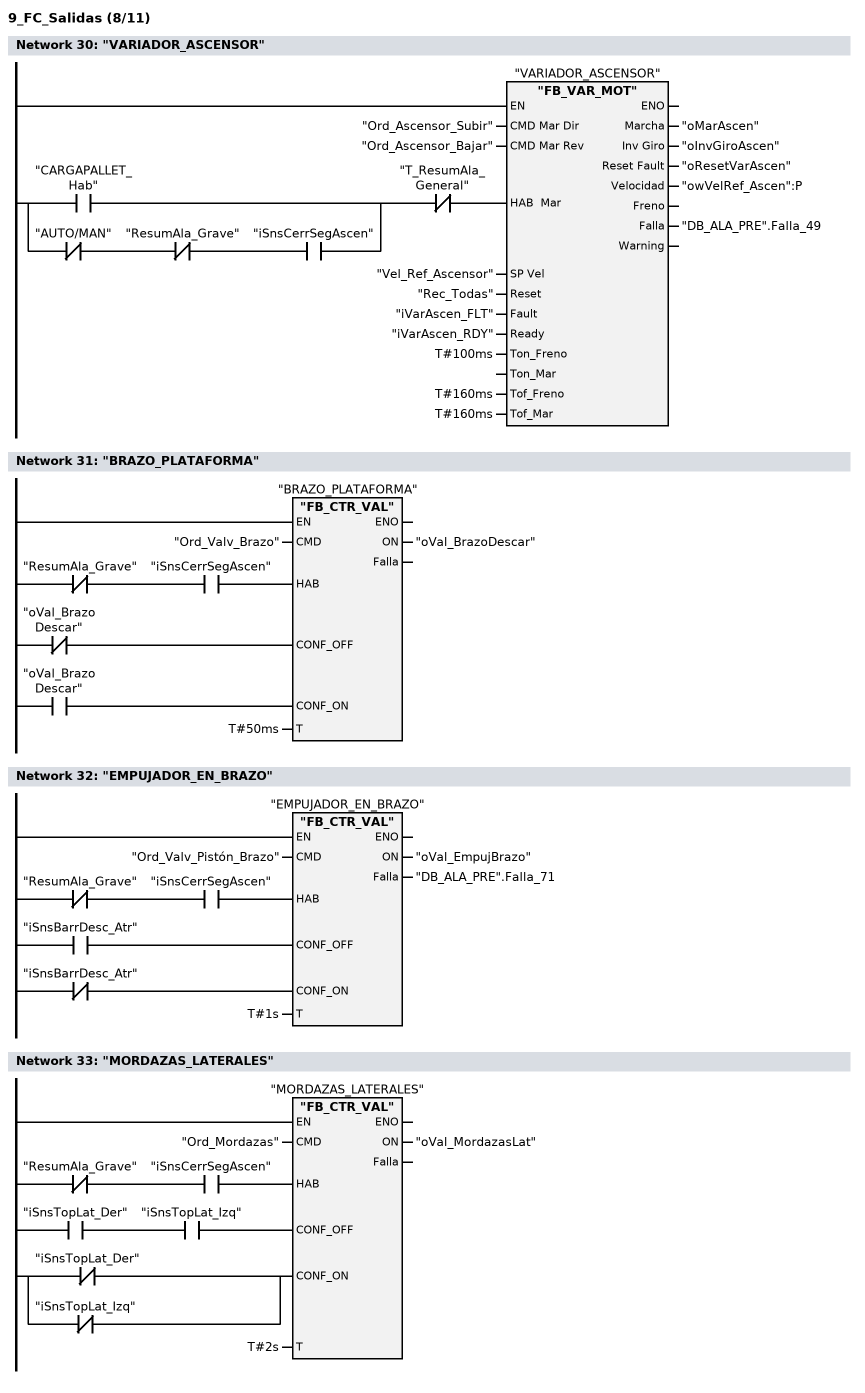
   RUNG wire#powerrail
      "VARIADOR_ASCENSOR"("HAB  Mar" := wire#w2, "CMD Mar Dir" := "Ord_Ascensor_Subir", "CMD Mar Rev" := "Ord_Ascensor_Bajar", "SP Vel" := "Vel_Ref_Ascensor", Reset := "Rec_Todas", Fault := "iVarAscen_FLT", Ready := "iVarAscen_RDY", Ton_Freno := T#100ms, Ton_Mar :=, Tof_Freno := T#160ms, Tof_Mar := T#160ms, Marcha => "oMarAscen", "Inv Giro" => "oInvGiroAscen", "Reset Fault" => "oResetVarAscen", Velocidad => "owVelRef_Ascen":P, Freno =>, Falla => "DB_ALA_PRE".Falla_49, Warning =>)
   END_RUNG
   RUNG wire#powerrail
      Contact( "CARGAPALLET_Hab" )
      wire#w1
      I_Contact( "T_ResumAla_General" )
   END_RUNG wire#w2
   RUNG wire#powerrail
      I_Contact( "AUTO/MAN" )
      I_Contact( "ResumAla_Grave" )
      Contact( "iSnsCerrSegAscen" )
   END_RUNG wire#w1
   // the same network as SCL:
   "VARIADOR_ASCENSOR"("CMD Mar Dir" := "Ord_Ascensor_Subir",   // "FB_VAR_MOT"
                       "CMD Mar Rev" := "Ord_Ascensor_Bajar",
                       "HAB  Mar" := ("CARGAPALLET_Hab" OR (NOT "AUTO/MAN" AND NOT "ResumAla_Grave" AND "iSnsCerrSegAscen")) AND NOT "T_ResumAla_General",
                       "SP Vel" := "Vel_Ref_Ascensor",
                       Reset := "Rec_Todas",
                       Fault := "iVarAscen_FLT",
                       Ready := "iVarAscen_RDY",
                       Ton_Freno := T#100ms,
                       Tof_Freno := T#160ms,
                       Tof_Mar := T#160ms,
                       Marcha => "oMarAscen",
                       "Inv Giro" => "oInvGiroAscen",
                       "Reset Fault" => "oResetVarAscen",
                       Velocidad => "owVelRef_Ascen":P,
                       Falla => "DB_ALA_PRE".Falla_49);
END_REGION

REGION Network 31: "BRAZO_PLATAFORMA"
   RUNG wire#powerrail
      "BRAZO_PLATAFORMA"(HAB := wire#w1, CONF_OFF := wire#w2, CONF_ON := wire#w3, CMD := "Ord_Valv_Brazo", T := T#50ms, ON => "oVal_BrazoDescar", Falla =>)
   END_RUNG
   RUNG wire#powerrail
      I_Contact( "ResumAla_Grave" )
      Contact( "iSnsCerrSegAscen" )
   END_RUNG wire#w1
   RUNG wire#powerrail
      I_Contact( "oVal_BrazoDescar" )
   END_RUNG wire#w2
   RUNG wire#powerrail
      Contact( "oVal_BrazoDescar" )
   END_RUNG wire#w3
   // the same network as SCL:
   "BRAZO_PLATAFORMA"(CMD := "Ord_Valv_Brazo",   // "FB_CTR_VAL"
                      HAB := NOT "ResumAla_Grave" AND "iSnsCerrSegAscen",
                      CONF_OFF := NOT "oVal_BrazoDescar",
                      CONF_ON := "oVal_BrazoDescar",
                      T := T#50ms,
                      ON => "oVal_BrazoDescar");
END_REGION

REGION Network 32: "EMPUJADOR_EN_BRAZO"
   RUNG wire#powerrail
      "EMPUJADOR_EN_BRAZO"(HAB := wire#w1, CONF_OFF := wire#w2, CONF_ON := wire#w3, CMD := "Ord_Valv_Pistón_Brazo", T := T#1s, ON => "oVal_EmpujBrazo", Falla => "DB_ALA_PRE".Falla_71)
   END_RUNG
   RUNG wire#powerrail
      I_Contact( "ResumAla_Grave" )
      Contact( "iSnsCerrSegAscen" )
   END_RUNG wire#w1
   RUNG wire#powerrail
      Contact( "iSnsBarrDesc_Atr" )
   END_RUNG wire#w2
   RUNG wire#powerrail
      I_Contact( "iSnsBarrDesc_Atr" )
   END_RUNG wire#w3
   // the same network as SCL:
   "EMPUJADOR_EN_BRAZO"(CMD := "Ord_Valv_Pistón_Brazo",   // "FB_CTR_VAL"
                        HAB := NOT "ResumAla_Grave" AND "iSnsCerrSegAscen",
                        CONF_OFF := "iSnsBarrDesc_Atr",
                        CONF_ON := NOT "iSnsBarrDesc_Atr",
                        T := T#1s,
                        ON => "oVal_EmpujBrazo",
                        Falla => "DB_ALA_PRE".Falla_71);
END_REGION

REGION Network 33: "MORDAZAS_LATERALES"
   RUNG wire#powerrail
      "MORDAZAS_LATERALES"(HAB := wire#w1, CONF_OFF := wire#w2, CONF_ON := wire#w3, CMD := "Ord_Mordazas", T := T#2s, ON => "oVal_MordazasLat", Falla =>)
   END_RUNG
   RUNG wire#powerrail
      I_Contact( "ResumAla_Grave" )
      Contact( "iSnsCerrSegAscen" )
   END_RUNG wire#w1
   RUNG wire#powerrail
      Contact( "iSnsTopLat_Der" )
      Contact( "iSnsTopLat_Izq" )
   END_RUNG wire#w2
   RUNG wire#powerrail
      I_Contact( "iSnsTopLat_Der" )
   END_RUNG wire#w3
   RUNG wire#powerrail
      I_Contact( "iSnsTopLat_Izq" )
   END_RUNG wire#w3
   // the same network as SCL:
   "MORDAZAS_LATERALES"(CMD := "Ord_Mordazas",   // "FB_CTR_VAL"
                        HAB := NOT "ResumAla_Grave" AND "iSnsCerrSegAscen",
                        CONF_OFF := "iSnsTopLat_Der" AND "iSnsTopLat_Izq",
                        CONF_ON := NOT "iSnsTopLat_Der" OR NOT "iSnsTopLat_Izq",
                        T := T#2s,
                        ON => "oVal_MordazasLat");
END_REGION

REGION Network 34: "MORDAZA_FINAL"
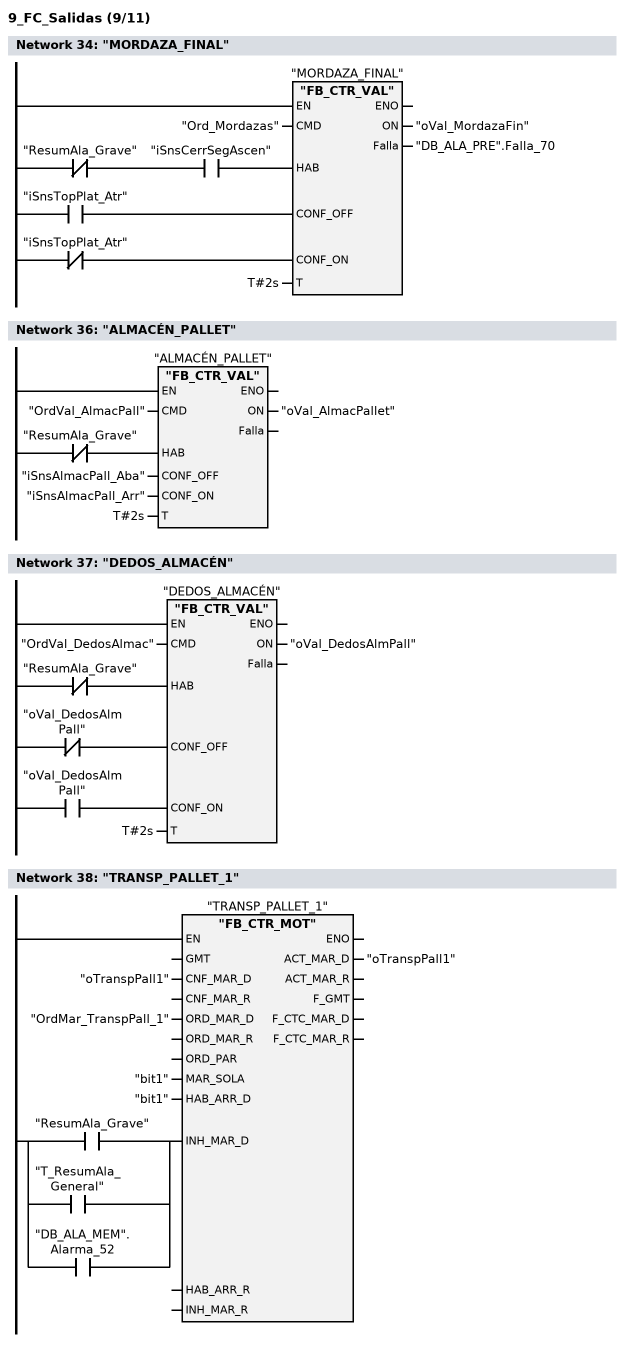
   RUNG wire#powerrail
      "MORDAZA_FINAL"(HAB := wire#w1, CONF_OFF := wire#w2, CONF_ON := wire#w3, CMD := "Ord_Mordazas", T := T#2s, ON => "oVal_MordazaFin", Falla => "DB_ALA_PRE".Falla_70)
   END_RUNG
   RUNG wire#powerrail
      I_Contact( "ResumAla_Grave" )
      Contact( "iSnsCerrSegAscen" )
   END_RUNG wire#w1
   RUNG wire#powerrail
      Contact( "iSnsTopPlat_Atr" )
   END_RUNG wire#w2
   RUNG wire#powerrail
      I_Contact( "iSnsTopPlat_Atr" )
   END_RUNG wire#w3
   // the same network as SCL:
   "MORDAZA_FINAL"(CMD := "Ord_Mordazas",   // "FB_CTR_VAL"
                   HAB := NOT "ResumAla_Grave" AND "iSnsCerrSegAscen",
                   CONF_OFF := "iSnsTopPlat_Atr",
                   CONF_ON := NOT "iSnsTopPlat_Atr",
                   T := T#2s,
                   ON => "oVal_MordazaFin",
                   Falla => "DB_ALA_PRE".Falla_70);
END_REGION

REGION Network 35: ----------------------------------------------------------------- TRANSPORTE DE PALLETS -----------------------------------------------------------------¬
END_REGION

REGION Network 36: "ALMACÉN_PALLET"
   RUNG wire#powerrail
      "ALMACÉN_PALLET"(HAB := wire#w1, CMD := "OrdVal_AlmacPall", CONF_OFF := "iSnsAlmacPall_Aba", CONF_ON := "iSnsAlmacPall_Arr", T := T#2s, ON => "oVal_AlmacPallet", Falla =>)
   END_RUNG
   RUNG wire#powerrail
      I_Contact( "ResumAla_Grave" )
   END_RUNG wire#w1
   // the same network as SCL:
   "ALMACÉN_PALLET"(CMD := "OrdVal_AlmacPall",   // "FB_CTR_VAL"
                    HAB := NOT "ResumAla_Grave",
                    CONF_OFF := "iSnsAlmacPall_Aba",
                    CONF_ON := "iSnsAlmacPall_Arr",
                    T := T#2s,
                    ON => "oVal_AlmacPallet");
END_REGION

REGION Network 37: "DEDOS_ALMACÉN"
   RUNG wire#powerrail
      "DEDOS_ALMACÉN"(HAB := wire#w1, CONF_OFF := wire#w2, CONF_ON := wire#w3, CMD := "OrdVal_DedosAlmac", T := T#2s, ON => "oVal_DedosAlmPall", Falla =>)
   END_RUNG
   RUNG wire#powerrail
      I_Contact( "ResumAla_Grave" )
   END_RUNG wire#w1
   RUNG wire#powerrail
      I_Contact( "oVal_DedosAlmPall" )
   END_RUNG wire#w2
   RUNG wire#powerrail
      Contact( "oVal_DedosAlmPall" )
   END_RUNG wire#w3
   // the same network as SCL:
   "DEDOS_ALMACÉN"(CMD := "OrdVal_DedosAlmac",   // "FB_CTR_VAL"
                   HAB := NOT "ResumAla_Grave",
                   CONF_OFF := NOT "oVal_DedosAlmPall",
                   CONF_ON := "oVal_DedosAlmPall",
                   T := T#2s,
                   ON => "oVal_DedosAlmPall");
END_REGION

REGION Network 38: "TRANSP_PALLET_1"
   RUNG wire#powerrail
      "TRANSP_PALLET_1"(INH_MAR_D := wire#w1, GMT :=, CNF_MAR_D := "oTranspPall1", CNF_MAR_R :=, ORD_MAR_D := "OrdMar_TranspPall_1", ORD_MAR_R :=, ORD_PAR :=, MAR_SOLA := "bit1", HAB_ARR_D := "bit1", HAB_ARR_R :=, INH_MAR_R :=, ACT_MAR_D => "oTranspPall1", ACT_MAR_R =>, F_GMT =>, F_CTC_MAR_D =>, F_CTC_MAR_R =>)
   END_RUNG
   RUNG wire#powerrail
      Contact( "ResumAla_Grave" )
   END_RUNG wire#w1
   RUNG wire#powerrail
      Contact( "T_ResumAla_General" )
   END_RUNG wire#w1
   RUNG wire#powerrail
      Contact( "DB_ALA_MEM".Alarma_52 )
   END_RUNG wire#w1
   // the same network as SCL:
   "TRANSP_PALLET_1"(CNF_MAR_D := "oTranspPall1",   // "FB_CTR_MOT"
                     ORD_MAR_D := "OrdMar_TranspPall_1",
                     MAR_SOLA := "bit1",
                     HAB_ARR_D := "bit1",
                     INH_MAR_D := "ResumAla_Grave" OR "T_ResumAla_General" OR "DB_ALA_MEM".Alarma_52,
                     ACT_MAR_D => "oTranspPall1");
END_REGION

REGION Network 39: "TRANSP_PALLET_2"
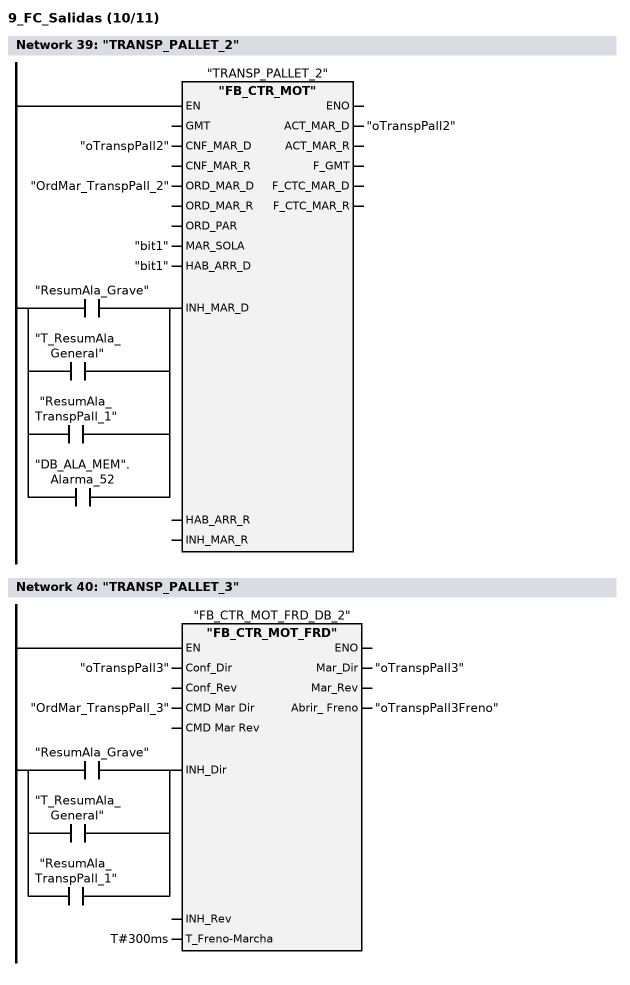
   RUNG wire#powerrail
      "TRANSP_PALLET_2"(INH_MAR_D := wire#w1, GMT :=, CNF_MAR_D := "oTranspPall2", CNF_MAR_R :=, ORD_MAR_D := "OrdMar_TranspPall_2", ORD_MAR_R :=, ORD_PAR :=, MAR_SOLA := "bit1", HAB_ARR_D := "bit1", HAB_ARR_R :=, INH_MAR_R :=, ACT_MAR_D => "oTranspPall2", ACT_MAR_R =>, F_GMT =>, F_CTC_MAR_D =>, F_CTC_MAR_R =>)
   END_RUNG
   RUNG wire#powerrail
      Contact( "ResumAla_Grave" )
   END_RUNG wire#w1
   RUNG wire#powerrail
      Contact( "T_ResumAla_General" )
   END_RUNG wire#w1
   RUNG wire#powerrail
      Contact( "ResumAla_TranspPall_1" )
   END_RUNG wire#w1
   RUNG wire#powerrail
      Contact( "DB_ALA_MEM".Alarma_52 )
   END_RUNG wire#w1
   // the same network as SCL:
   "TRANSP_PALLET_2"(CNF_MAR_D := "oTranspPall2",   // "FB_CTR_MOT"
                     ORD_MAR_D := "OrdMar_TranspPall_2",
                     MAR_SOLA := "bit1",
                     HAB_ARR_D := "bit1",
                     INH_MAR_D := "ResumAla_Grave" OR "T_ResumAla_General" OR "ResumAla_TranspPall_1" OR "DB_ALA_MEM".Alarma_52,
                     ACT_MAR_D => "oTranspPall2");
END_REGION

REGION Network 40: "TRANSP_PALLET_3"
   RUNG wire#powerrail
      "FB_CTR_MOT_FRD_DB_2"(INH_Dir := wire#w1, Conf_Dir := "oTranspPall3", Conf_Rev :=, "CMD Mar Dir" := "OrdMar_TranspPall_3", "CMD Mar Rev" :=, INH_Rev :=, "T_Freno-Marcha" := T#300ms, Mar_Dir => "oTranspPall3", Mar_Rev =>, "Abrir_ Freno" => "oTranspPall3Freno")
   END_RUNG
   RUNG wire#powerrail
      Contact( "ResumAla_Grave" )
   END_RUNG wire#w1
   RUNG wire#powerrail
      Contact( "T_ResumAla_General" )
   END_RUNG wire#w1
   RUNG wire#powerrail
      Contact( "ResumAla_TranspPall_1" )
   END_RUNG wire#w1
   // the same network as SCL:
   "FB_CTR_MOT_FRD_DB_2"(Conf_Dir := "oTranspPall3",   // "FB_CTR_MOT_FRD"
                         "CMD Mar Dir" := "OrdMar_TranspPall_3",
                         INH_Dir := "ResumAla_Grave" OR "T_ResumAla_General" OR "ResumAla_TranspPall_1",
                         "T_Freno-Marcha" := T#300ms,
                         Mar_Dir => "oTranspPall3",
                         "Abrir_ Freno" => "oTranspPall3Freno");
END_REGION

REGION Network 41: "TRANSP_PALLET_4"
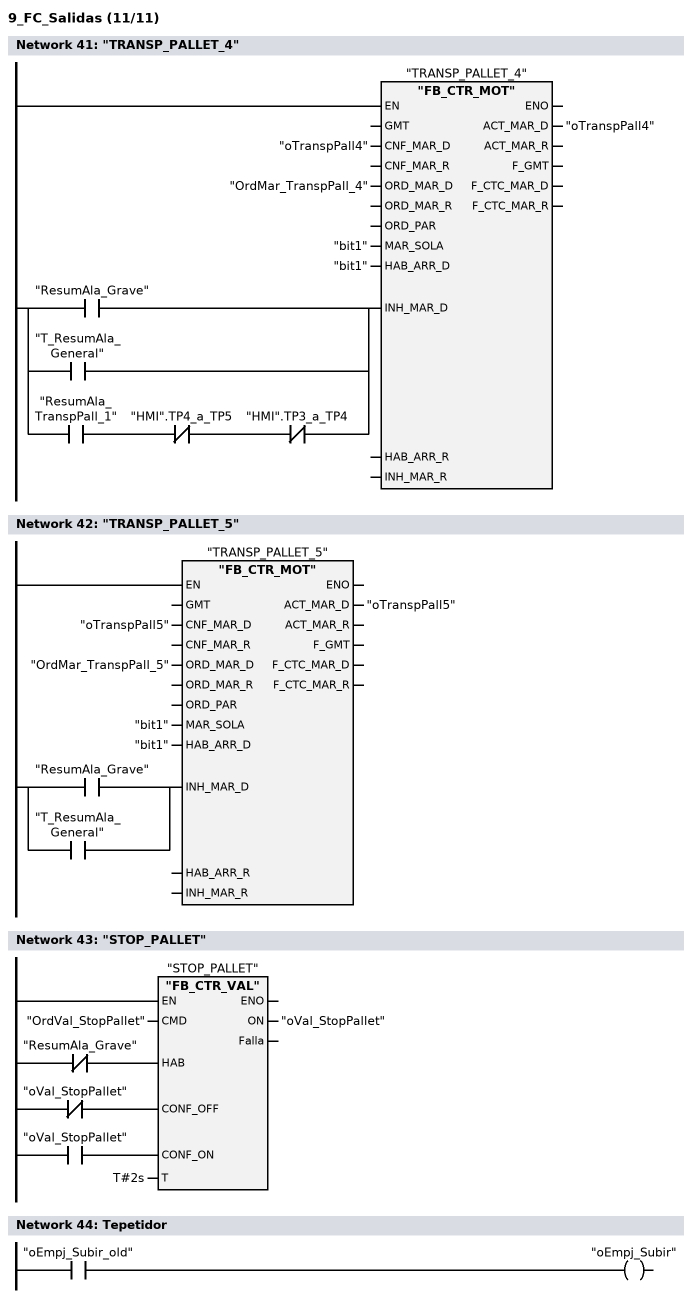
   RUNG wire#powerrail
      "TRANSP_PALLET_4"(INH_MAR_D := wire#w1, GMT :=, CNF_MAR_D := "oTranspPall4", CNF_MAR_R :=, ORD_MAR_D := "OrdMar_TranspPall_4", ORD_MAR_R :=, ORD_PAR :=, MAR_SOLA := "bit1", HAB_ARR_D := "bit1", HAB_ARR_R :=, INH_MAR_R :=, ACT_MAR_D => "oTranspPall4", ACT_MAR_R =>, F_GMT =>, F_CTC_MAR_D =>, F_CTC_MAR_R =>)
   END_RUNG
   RUNG wire#powerrail
      Contact( "ResumAla_Grave" )
   END_RUNG wire#w1
   RUNG wire#powerrail
      Contact( "T_ResumAla_General" )
   END_RUNG wire#w1
   RUNG wire#powerrail
      Contact( "ResumAla_TranspPall_1" )
      I_Contact( "HMI".TP4_a_TP5 )
      I_Contact( "HMI".TP3_a_TP4 )
   END_RUNG wire#w1
   // the same network as SCL:
   "TRANSP_PALLET_4"(CNF_MAR_D := "oTranspPall4",   // "FB_CTR_MOT"
                     ORD_MAR_D := "OrdMar_TranspPall_4",
                     MAR_SOLA := "bit1",
                     HAB_ARR_D := "bit1",
                     INH_MAR_D := "ResumAla_Grave" OR "T_ResumAla_General" OR ("ResumAla_TranspPall_1" AND NOT "HMI".TP4_a_TP5 AND NOT "HMI".TP3_a_TP4),
                     ACT_MAR_D => "oTranspPall4");
END_REGION

REGION Network 42: "TRANSP_PALLET_5"
   RUNG wire#powerrail
      "TRANSP_PALLET_5"(INH_MAR_D := wire#w1, GMT :=, CNF_MAR_D := "oTranspPall5", CNF_MAR_R :=, ORD_MAR_D := "OrdMar_TranspPall_5", ORD_MAR_R :=, ORD_PAR :=, MAR_SOLA := "bit1", HAB_ARR_D := "bit1", HAB_ARR_R :=, INH_MAR_R :=, ACT_MAR_D => "oTranspPall5", ACT_MAR_R =>, F_GMT =>, F_CTC_MAR_D =>, F_CTC_MAR_R =>)
   END_RUNG
   RUNG wire#powerrail
      Contact( "ResumAla_Grave" )
   END_RUNG wire#w1
   RUNG wire#powerrail
      Contact( "T_ResumAla_General" )
   END_RUNG wire#w1
   // the same network as SCL:
   "TRANSP_PALLET_5"(CNF_MAR_D := "oTranspPall5",   // "FB_CTR_MOT"
                     ORD_MAR_D := "OrdMar_TranspPall_5",
                     MAR_SOLA := "bit1",
                     HAB_ARR_D := "bit1",
                     INH_MAR_D := "ResumAla_Grave" OR "T_ResumAla_General",
                     ACT_MAR_D => "oTranspPall5");
END_REGION

REGION Network 43: "STOP_PALLET"
   RUNG wire#powerrail
      "STOP_PALLET"(HAB := wire#w1, CONF_OFF := wire#w2, CONF_ON := wire#w3, CMD := "OrdVal_StopPallet", T := T#2s, ON => "oVal_StopPallet", Falla =>)
   END_RUNG
   RUNG wire#powerrail
      I_Contact( "ResumAla_Grave" )
   END_RUNG wire#w1
   RUNG wire#powerrail
      I_Contact( "oVal_StopPallet" )
   END_RUNG wire#w2
   RUNG wire#powerrail
      Contact( "oVal_StopPallet" )
   END_RUNG wire#w3
   // the same network as SCL:
   "STOP_PALLET"(CMD := "OrdVal_StopPallet",   // "FB_CTR_VAL"
                 HAB := NOT "ResumAla_Grave",
                 CONF_OFF := NOT "oVal_StopPallet",
                 CONF_ON := "oVal_StopPallet",
                 T := T#2s,
                 ON => "oVal_StopPallet");
END_REGION

REGION Network 44: Tepetidor
   RUNG wire#powerrail
      Contact( "oEmpj_Subir_old" )
      Coil( "oEmpj_Subir" )
   END_RUNG
   // the same network as SCL:
   "oEmpj_Subir" := "oEmpj_Subir_old";
END_REGION
END_FUNCTION

FUNCTION "4_FC_Dosificador" : Void   // FC11, LAD
{ S7_Optimized_Access := 'FALSE' }
VERSION : 0.1
BEGIN

REGION Network 1: ESTADO ACTIVO
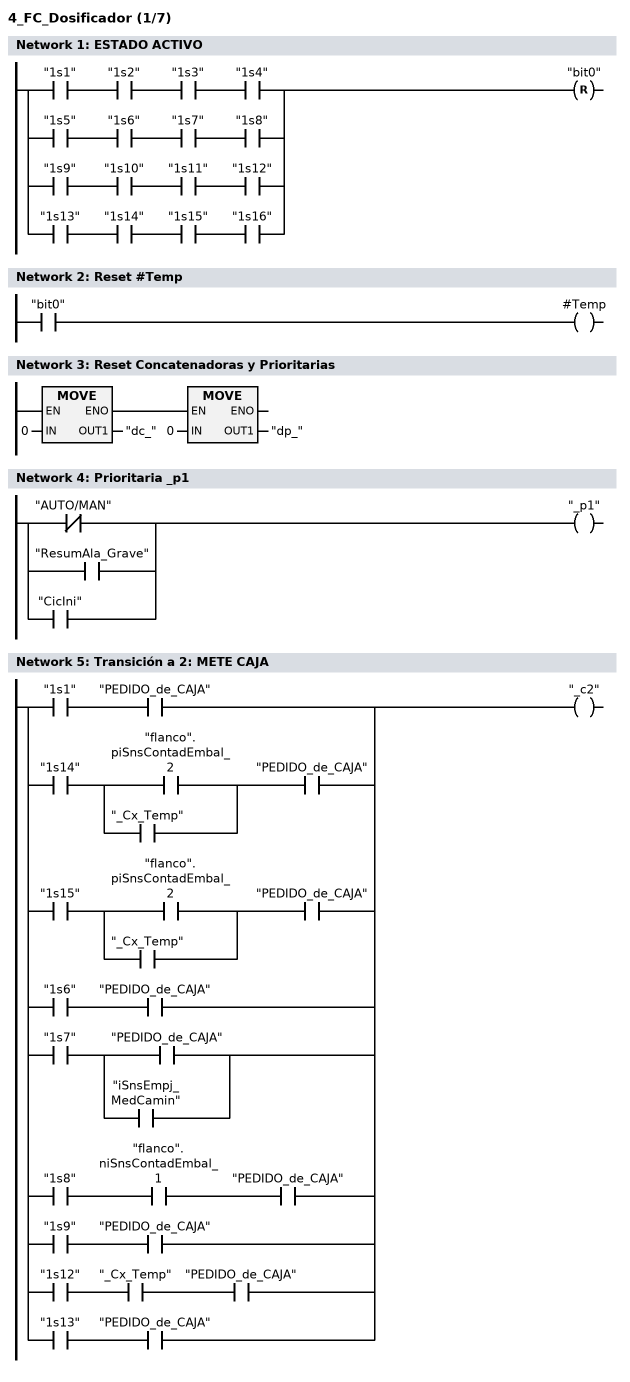
   RUNG wire#powerrail
      Contact( "1s1" )
      Contact( "1s2" )
      Contact( "1s3" )
      Contact( "1s4" )
      wire#w1
      R_Coil( "bit0" )
   END_RUNG
   RUNG wire#powerrail
      Contact( "1s5" )
      Contact( "1s6" )
      Contact( "1s7" )
      Contact( "1s8" )
   END_RUNG wire#w1
   RUNG wire#powerrail
      Contact( "1s9" )
      Contact( "1s10" )
      Contact( "1s11" )
      Contact( "1s12" )
   END_RUNG wire#w1
   RUNG wire#powerrail
      Contact( "1s13" )
      Contact( "1s14" )
      Contact( "1s15" )
      Contact( "1s16" )
   END_RUNG wire#w1
   // the same network as SCL:
   IF ("1s1" AND "1s2" AND "1s3" AND "1s4") OR ("1s5" AND "1s6" AND "1s7" AND "1s8") OR ("1s9" AND "1s10" AND "1s11" AND "1s12") OR ("1s13" AND "1s14" AND "1s15" AND "1s16") THEN
       "bit0" := FALSE;
   END_IF;
END_REGION

REGION Network 2: Reset #Temp
   RUNG wire#powerrail
      Contact( "bit0" )
      Coil( #Temp )
   END_RUNG
   // the same network as SCL:
   #Temp := "bit0";
END_REGION

REGION Network 3: Reset Concatenadoras y Prioritarias
   RUNG wire#powerrail
      { S7_GenerateENO := "TRUE" } Move(in := 0, out1 => "dc_")
      { S7_GenerateENO := "TRUE" } Move(in := 0, out1 => "dp_")
   END_RUNG
   // the same network as SCL:
   // ENO of a box is taken as its EN; it also drops when the box reports an error
   "dc_" := 0;
   "dp_" := 0;
END_REGION

REGION Network 4: Prioritaria _p1
   RUNG wire#powerrail
      I_Contact( "AUTO/MAN" )
      wire#w1
      Coil( "_p1" )
   END_RUNG
   RUNG wire#powerrail
      Contact( "ResumAla_Grave" )
   END_RUNG wire#w1
   RUNG wire#powerrail
      Contact( "CicIni" )
   END_RUNG wire#w1
   // the same network as SCL:
   "_p1" := NOT "AUTO/MAN" OR "ResumAla_Grave" OR "CicIni";
END_REGION

REGION Network 5: Transición a 2: METE CAJA
   RUNG wire#powerrail
      Contact( "1s1" )
      Contact( "PEDIDO_de_CAJA" )
      wire#w1
      Coil( "_c2" )
   END_RUNG
   RUNG wire#powerrail
      Contact( "1s14" )
      wire#w2
      Contact( "flanco".piSnsContadEmbal_2 )
      wire#w3
      Contact( "PEDIDO_de_CAJA" )
   END_RUNG wire#w1
   RUNG wire#w2
      Contact( "_Cx_Temp" )
   END_RUNG wire#w3
   RUNG wire#powerrail
      Contact( "1s15" )
      wire#w4
      Contact( "flanco".piSnsContadEmbal_2 )
      wire#w5
      Contact( "PEDIDO_de_CAJA" )
   END_RUNG wire#w1
   RUNG wire#w4
      Contact( "_Cx_Temp" )
   END_RUNG wire#w5
   RUNG wire#powerrail
      Contact( "1s6" )
      Contact( "PEDIDO_de_CAJA" )
   END_RUNG wire#w1
   RUNG wire#powerrail
      Contact( "1s7" )
      wire#w6
      Contact( "PEDIDO_de_CAJA" )
   END_RUNG wire#w1
   RUNG wire#w6
      Contact( "iSnsEmpj_MedCamin" )
   END_RUNG wire#w1
   RUNG wire#powerrail
      Contact( "1s8" )
      Contact( "flanco".niSnsContadEmbal_1 )
      Contact( "PEDIDO_de_CAJA" )
   END_RUNG wire#w1
   RUNG wire#powerrail
      Contact( "1s9" )
      Contact( "PEDIDO_de_CAJA" )
   END_RUNG wire#w1
   RUNG wire#powerrail
      Contact( "1s12" )
      Contact( "_Cx_Temp" )
      Contact( "PEDIDO_de_CAJA" )
   END_RUNG wire#w1
   RUNG wire#powerrail
      Contact( "1s13" )
      Contact( "PEDIDO_de_CAJA" )
   END_RUNG wire#w1
   // the same network as SCL:
   "_c2" := ("1s1" AND "PEDIDO_de_CAJA") OR ("1s14" AND ("flanco".piSnsContadEmbal_2 OR "_Cx_Temp") AND "PEDIDO_de_CAJA") OR ("1s15" AND ("flanco".piSnsContadEmbal_2 OR "_Cx_Temp") AND "PEDIDO_de_CAJA") OR ("1s6" AND "PEDIDO_de_CAJA") OR ("1s7" AND ("PEDIDO_de_CAJA" OR "iSnsEmpj_MedCamin")) OR ("1s8" AND "flanco".niSnsContadEmbal_1 AND "PEDIDO_de_CAJA") OR ("1s9" AND "PEDIDO_de_CAJA") OR ("1s12" AND "_Cx_Temp" AND "PEDIDO_de_CAJA") OR ("1s13" AND "PEDIDO_de_CAJA");
END_REGION

REGION Network 6: Transición a 3: FIGURA H
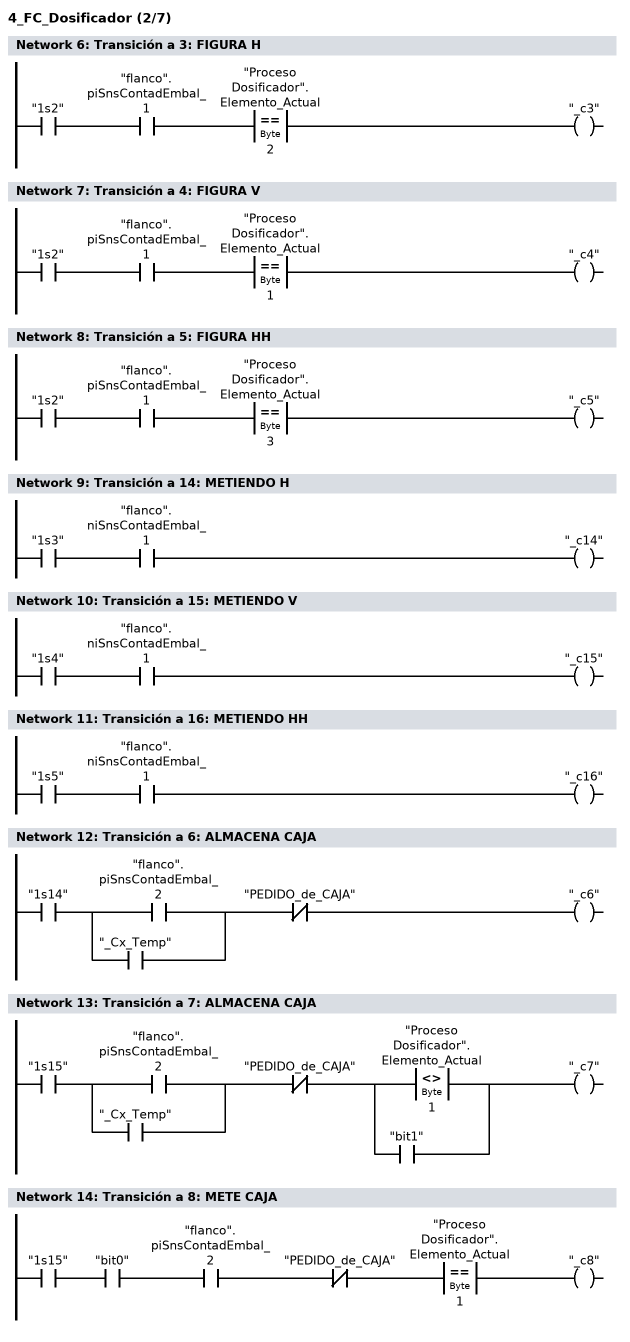
   RUNG wire#powerrail
      Contact( "1s2" )
      Contact( "flanco".piSnsContadEmbal_1 )
      { S7_Templates := "SrcType := Byte" } EQ_Contact(in1 := "Proceso Dosificador".Elemento_Actual, in2 := 2)
      Coil( "_c3" )
   END_RUNG
   // the same network as SCL:
   "_c3" := "1s2" AND "flanco".piSnsContadEmbal_1 AND ("Proceso Dosificador".Elemento_Actual = 2);
END_REGION

REGION Network 7: Transición a 4: FIGURA V
   RUNG wire#powerrail
      Contact( "1s2" )
      Contact( "flanco".piSnsContadEmbal_1 )
      { S7_Templates := "SrcType := Byte" } EQ_Contact(in1 := "Proceso Dosificador".Elemento_Actual, in2 := 1)
      Coil( "_c4" )
   END_RUNG
   // the same network as SCL:
   "_c4" := "1s2" AND "flanco".piSnsContadEmbal_1 AND ("Proceso Dosificador".Elemento_Actual = 1);
END_REGION

REGION Network 8: Transición a 5: FIGURA HH
   RUNG wire#powerrail
      Contact( "1s2" )
      Contact( "flanco".piSnsContadEmbal_1 )
      { S7_Templates := "SrcType := Byte" } EQ_Contact(in1 := "Proceso Dosificador".Elemento_Actual, in2 := 3)
      Coil( "_c5" )
   END_RUNG
   // the same network as SCL:
   "_c5" := "1s2" AND "flanco".piSnsContadEmbal_1 AND ("Proceso Dosificador".Elemento_Actual = 3);
END_REGION

REGION Network 9: Transición a 14: METIENDO H
   RUNG wire#powerrail
      Contact( "1s3" )
      Contact( "flanco".niSnsContadEmbal_1 )
      Coil( "_c14" )
   END_RUNG
   // the same network as SCL:
   "_c14" := "1s3" AND "flanco".niSnsContadEmbal_1;
END_REGION

REGION Network 10: Transición a 15: METIENDO V
   RUNG wire#powerrail
      Contact( "1s4" )
      Contact( "flanco".niSnsContadEmbal_1 )
      Coil( "_c15" )
   END_RUNG
   // the same network as SCL:
   "_c15" := "1s4" AND "flanco".niSnsContadEmbal_1;
END_REGION

REGION Network 11: Transición a 16: METIENDO HH
   RUNG wire#powerrail
      Contact( "1s5" )
      Contact( "flanco".niSnsContadEmbal_1 )
      Coil( "_c16" )
   END_RUNG
   // the same network as SCL:
   "_c16" := "1s5" AND "flanco".niSnsContadEmbal_1;
END_REGION

REGION Network 12: Transición a 6: ALMACENA CAJA
   RUNG wire#powerrail
      Contact( "1s14" )
      wire#w1
      Contact( "flanco".piSnsContadEmbal_2 )
      wire#w2
      I_Contact( "PEDIDO_de_CAJA" )
      Coil( "_c6" )
   END_RUNG
   RUNG wire#w1
      Contact( "_Cx_Temp" )
   END_RUNG wire#w2
   // the same network as SCL:
   "_c6" := "1s14" AND ("flanco".piSnsContadEmbal_2 OR "_Cx_Temp") AND NOT "PEDIDO_de_CAJA";
END_REGION

REGION Network 13: Transición a 7: ALMACENA CAJA
   RUNG wire#powerrail
      Contact( "1s15" )
      wire#w1
      Contact( "flanco".piSnsContadEmbal_2 )
      wire#w2
      I_Contact( "PEDIDO_de_CAJA" )
      wire#w3
      { S7_Templates := "SrcType := Byte" } NE_Contact(in1 := "Proceso Dosificador".Elemento_Actual, in2 := 1)
      wire#w4
      Coil( "_c7" )
   END_RUNG
   RUNG wire#w1
      Contact( "_Cx_Temp" )
   END_RUNG wire#w2
   RUNG wire#w3
      Contact( "bit1" )
   END_RUNG wire#w4
   // the same network as SCL:
   "_c7" := "1s15" AND ("flanco".piSnsContadEmbal_2 OR "_Cx_Temp") AND NOT "PEDIDO_de_CAJA" AND (("Proceso Dosificador".Elemento_Actual <> 1) OR "bit1");
END_REGION

REGION Network 14: Transición a 8: METE CAJA
   RUNG wire#powerrail
      Contact( "1s15" )
      Contact( "bit0" )
      Contact( "flanco".piSnsContadEmbal_2 )
      I_Contact( "PEDIDO_de_CAJA" )
      { S7_Templates := "SrcType := Byte" } EQ_Contact(in1 := "Proceso Dosificador".Elemento_Actual, in2 := 1)
      Coil( "_c8" )
   END_RUNG
   // the same network as SCL:
   "_c8" := "1s15" AND "bit0" AND "flanco".piSnsContadEmbal_2 AND NOT "PEDIDO_de_CAJA" AND ("Proceso Dosificador".Elemento_Actual = 1);
END_REGION

REGION Network 15: Transición a 9: ALMACENA CAJA
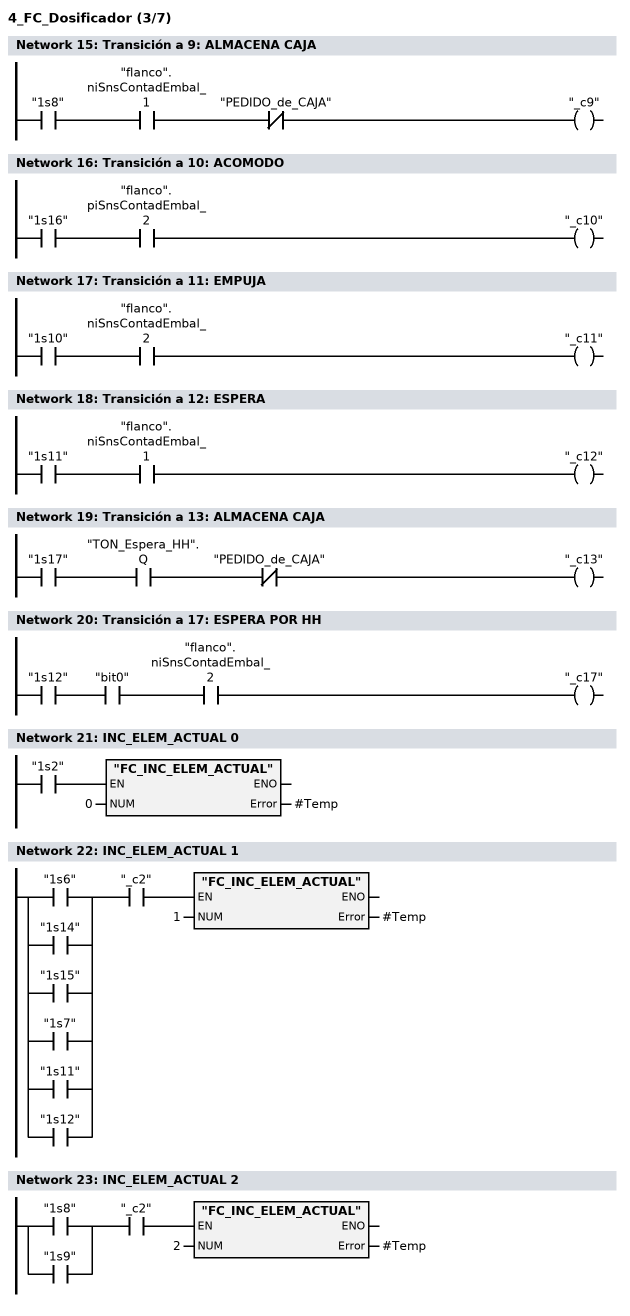
   RUNG wire#powerrail
      Contact( "1s8" )
      Contact( "flanco".niSnsContadEmbal_1 )
      I_Contact( "PEDIDO_de_CAJA" )
      Coil( "_c9" )
   END_RUNG
   // the same network as SCL:
   "_c9" := "1s8" AND "flanco".niSnsContadEmbal_1 AND NOT "PEDIDO_de_CAJA";
END_REGION

REGION Network 16: Transición a 10: ACOMODO
   RUNG wire#powerrail
      Contact( "1s16" )
      Contact( "flanco".piSnsContadEmbal_2 )
      Coil( "_c10" )
   END_RUNG
   // the same network as SCL:
   "_c10" := "1s16" AND "flanco".piSnsContadEmbal_2;
END_REGION

REGION Network 17: Transición a 11: EMPUJA
   RUNG wire#powerrail
      Contact( "1s10" )
      Contact( "flanco".niSnsContadEmbal_2 )
      Coil( "_c11" )
   END_RUNG
   // the same network as SCL:
   "_c11" := "1s10" AND "flanco".niSnsContadEmbal_2;
END_REGION

REGION Network 18: Transición a 12: ESPERA
   RUNG wire#powerrail
      Contact( "1s11" )
      Contact( "flanco".niSnsContadEmbal_1 )
      Coil( "_c12" )
   END_RUNG
   // the same network as SCL:
   "_c12" := "1s11" AND "flanco".niSnsContadEmbal_1;
END_REGION

REGION Network 19: Transición a 13: ALMACENA CAJA
   RUNG wire#powerrail
      Contact( "1s17" )
      Contact( "TON_Espera_HH".Q )
      I_Contact( "PEDIDO_de_CAJA" )
      Coil( "_c13" )
   END_RUNG
   // the same network as SCL:
   "_c13" := "1s17" AND "TON_Espera_HH".Q AND NOT "PEDIDO_de_CAJA";
END_REGION

REGION Network 20: Transición a 17: ESPERA POR HH
   RUNG wire#powerrail
      Contact( "1s12" )
      Contact( "bit0" )
      Contact( "flanco".niSnsContadEmbal_2 )
      Coil( "_c17" )
   END_RUNG
   // the same network as SCL:
   "_c17" := "1s12" AND "bit0" AND "flanco".niSnsContadEmbal_2;
END_REGION

REGION Network 21: INC_ELEM_ACTUAL 0
   RUNG wire#powerrail
      Contact( "1s2" )
      "FC_INC_ELEM_ACTUAL"(NUM := 0, Error => #Temp)
   END_RUNG
   // the same network as SCL:
   IF "1s2" THEN "FC_INC_ELEM_ACTUAL"(NUM := 0, Error => #Temp); END_IF;
END_REGION

REGION Network 22: INC_ELEM_ACTUAL 1
   RUNG wire#powerrail
      Contact( "1s6" )
      wire#w1
      Contact( "_c2" )
      "FC_INC_ELEM_ACTUAL"(NUM := 1, Error => #Temp)
   END_RUNG
   RUNG wire#powerrail
      Contact( "1s14" )
   END_RUNG wire#w1
   RUNG wire#powerrail
      Contact( "1s15" )
   END_RUNG wire#w1
   RUNG wire#powerrail
      Contact( "1s7" )
   END_RUNG wire#w1
   RUNG wire#powerrail
      Contact( "1s11" )
   END_RUNG wire#w1
   RUNG wire#powerrail
      Contact( "1s12" )
   END_RUNG wire#w1
   // the same network as SCL:
   IF ("1s6" OR "1s14" OR "1s15" OR "1s7" OR "1s11" OR "1s12") AND "_c2" THEN
       "FC_INC_ELEM_ACTUAL"(NUM := 1, Error => #Temp);
   END_IF;
END_REGION

REGION Network 23: INC_ELEM_ACTUAL 2
   RUNG wire#powerrail
      Contact( "1s8" )
      wire#w1
      Contact( "_c2" )
      "FC_INC_ELEM_ACTUAL"(NUM := 2, Error => #Temp)
   END_RUNG
   RUNG wire#powerrail
      Contact( "1s9" )
   END_RUNG wire#w1
   // the same network as SCL:
   IF ("1s8" OR "1s9") AND "_c2" THEN "FC_INC_ELEM_ACTUAL"(NUM := 2, Error => #Temp); END_IF;
END_REGION

REGION Network 24: Error Programación
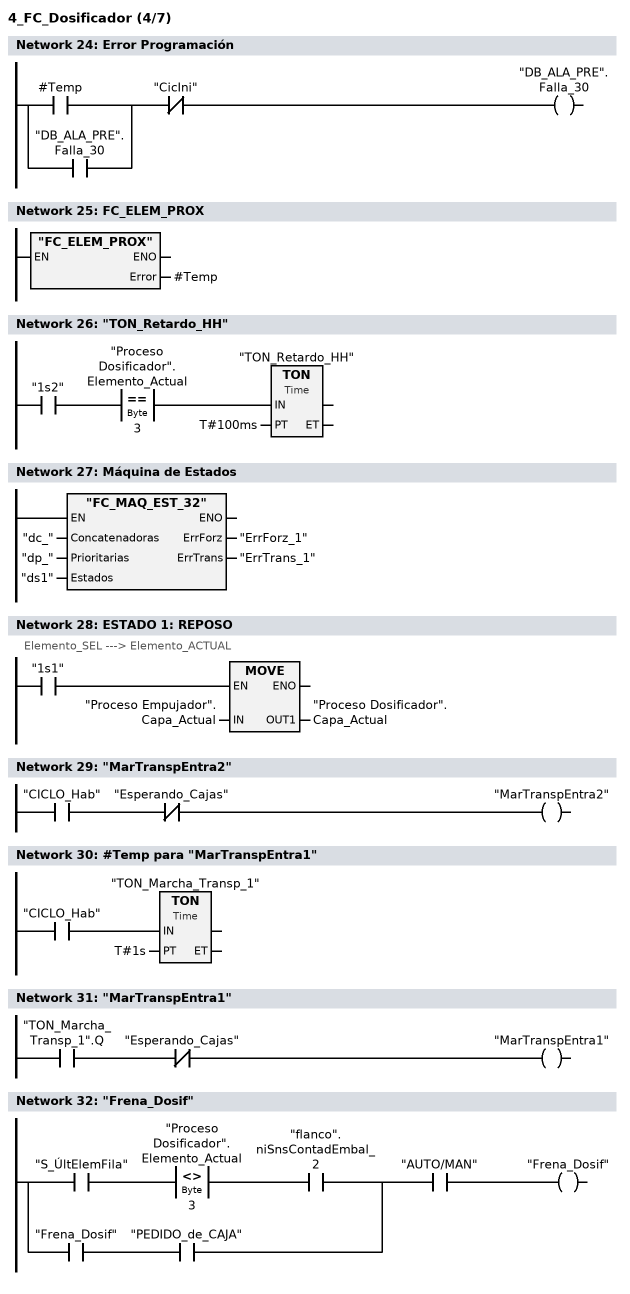
   RUNG wire#powerrail
      Contact( #Temp )
      wire#w1
      I_Contact( "CicIni" )
      Coil( "DB_ALA_PRE".Falla_30 )
   END_RUNG
   RUNG wire#powerrail
      Contact( "DB_ALA_PRE".Falla_30 )
   END_RUNG wire#w1
   // the same network as SCL:
   "DB_ALA_PRE".Falla_30 := (#Temp OR "DB_ALA_PRE".Falla_30) AND NOT "CicIni";
END_REGION

REGION Network 25: FC_ELEM_PROX
   RUNG wire#powerrail
      "FC_ELEM_PROX"(Error => #Temp)
   END_RUNG
   // the same network as SCL:
   "FC_ELEM_PROX"(Error => #Temp);
END_REGION

REGION Network 26: "TON_Retardo_HH"
   "TON_Retardo_HH".TON(in := "1s2" AND ("Proceso Dosificador".Elemento_Actual = 3), pt := T#100ms);
END_REGION

REGION Network 27: Máquina de Estados
   RUNG wire#powerrail
      "FC_MAQ_EST_32"(Concatenadoras := "dc_", Prioritarias := "dp_", Estados := "ds1", ErrForz => "ErrForz_1", ErrTrans => "ErrTrans_1")
   END_RUNG
   // the same network as SCL:
   "FC_MAQ_EST_32"(Concatenadoras := "dc_",
                   Prioritarias := "dp_",
                   Estados := "ds1",
                   ErrForz => "ErrForz_1",
                   ErrTrans => "ErrTrans_1");
END_REGION

REGION Network 28: ESTADO 1: REPOSO
   // Elemento_SEL ---> Elemento_ACTUAL
   RUNG wire#powerrail
      Contact( "1s1" )
      { S7_GenerateENO := "TRUE" } Move(in := "Proceso Empujador".Capa_Actual, out1 => "Proceso Dosificador".Capa_Actual)
   END_RUNG
   // the same network as SCL:
   IF "1s1" THEN "Proceso Dosificador".Capa_Actual := "Proceso Empujador".Capa_Actual; END_IF;
END_REGION

REGION Network 29: "MarTranspEntra2"
   RUNG wire#powerrail
      Contact( "CICLO_Hab" )
      I_Contact( "Esperando_Cajas" )
      Coil( "MarTranspEntra2" )
   END_RUNG
   // the same network as SCL:
   "MarTranspEntra2" := "CICLO_Hab" AND NOT "Esperando_Cajas";
END_REGION

REGION Network 30: #Temp para "MarTranspEntra1"
   "TON_Marcha_Transp_1".TON(in := "CICLO_Hab", pt := T#1s);
END_REGION

REGION Network 31: "MarTranspEntra1"
   RUNG wire#powerrail
      Contact( "TON_Marcha_Transp_1".Q )
      I_Contact( "Esperando_Cajas" )
      Coil( "MarTranspEntra1" )
   END_RUNG
   // the same network as SCL:
   "MarTranspEntra1" := "TON_Marcha_Transp_1".Q AND NOT "Esperando_Cajas";
END_REGION
